   "20_TANKS_IP_DATA_RIO_07_FIRST_TANK_USD_FLOW" : Real = PLC "20_TANKS_IP_DATA".RIO_07.FIRST_TANK.USD_FLOW, 1 s
   "20_TANKS_IP_DATA_RIO_07_FIRST_TANK_MBG_FLOW" : Real = PLC "20_TANKS_IP_DATA".RIO_07.FIRST_TANK.MBG_FLOW, 1 s
   "504_Tank Grouping_DB2020_RUN TANK 14" : Bool = PLC "504_Tank Grouping_DB2020"."RUN TANK 14", 1 s
   "504_Tank Grouping_DB2020_RUN TANK 6" : Bool = PLC "504_Tank Grouping_DB2020"."RUN TANK 6", 1 s
   "504_Tank Grouping_DB2020_RUN TANK 8" : Bool = PLC "504_Tank Grouping_DB2020"."RUN TANK 8", 1 s
   "504_Tank Grouping_DB2020_RUN TANK 9" : Bool = PLC "504_Tank Grouping_DB2020"."RUN TANK 9", 1 s
   "504_Tank Grouping_DB2020_RUN TANK 10" : Bool = PLC "504_Tank Grouping_DB2020"."RUN TANK 10", 1 s
   "504_Tank Grouping_DB2020_RUN TANK 11" : Bool = PLC "504_Tank Grouping_DB2020"."RUN TANK 11", 1 s
   "504_Tank Grouping_DB2020_RUN TANK 12" : Bool = PLC "504_Tank Grouping_DB2020"."RUN TANK 12", 1 s
   "504_Tank Grouping_DB2020_RUN TANK 13" : Bool = PLC "504_Tank Grouping_DB2020"."RUN TANK 13", 1 s
   "504_Tank Grouping_DB2020_Sequence Time m Offset" : Time = PLC "504_Tank Grouping_DB2020"."Sequence Time m Offset", 1 s
   "20_TANKS_IP_DATA_RIO_01_FIRST_TANK_TANKS_PRESS" : Real = PLC "20_TANKS_IP_DATA".RIO_01.FIRST_TANK.TANKS_PRESS, 1 s
   "20_TANKS_IP_DATA_RIO_01_FIRST_TANK_BWT_LEVEL" : Real = PLC "20_TANKS_IP_DATA".RIO_01.FIRST_TANK.BWT_LEVEL, 1 s
   "20_TANKS_IP_DATA_RIO_01_FIRST_TANK_BWT_PH" : Real = PLC "20_TANKS_IP_DATA".RIO_01.FIRST_TANK.BWT_PH, 1 s
   "20_TANKS_IP_DATA_RIO_01_FIRST_TANK_BWT_DO" : Real = PLC "20_TANKS_IP_DATA".RIO_01.FIRST_TANK.BWT_DO, 1 s
   "20_TANKS_IP_DATA_RIO_01_FIRST_TANK_BWT_TEMP" : Real = PLC "20_TANKS_IP_DATA".RIO_01.FIRST_TANK.BWT_TEMP, 1 s
   "504_Tank Grouping_DB2020_Tank1 Min Time_ET" : Time = PLC "504_Tank Grouping_DB2020"."Tank1 Min Time".ET, 1 s
   "504_Tank Grouping_DB2020_Tank2 Min Time_ET" : Time = PLC "504_Tank Grouping_DB2020"."Tank2 Min Time".ET, 1 s
   "20_TANKS_IP_DATA_RIO_01_SECOND_TANK_TANKS_PRESS" : Real = PLC "20_TANKS_IP_DATA".RIO_01.SECOND_TANK.TANKS_PRESS, 1 s
   "20_TANKS_IP_DATA_RIO_01_SECOND_TANK_BWT_LEVEL" : Real = PLC "20_TANKS_IP_DATA".RIO_01.SECOND_TANK.BWT_LEVEL, 1 s
   "20_TANKS_IP_DATA_RIO_01_SECOND_TANK_BWT_PH" : Real = PLC "20_TANKS_IP_DATA".RIO_01.SECOND_TANK.BWT_PH, 1 s
   "20_TANKS_IP_DATA_RIO_01_SECOND_TANK_BWT_DO" : Real = PLC "20_TANKS_IP_DATA".RIO_01.SECOND_TANK.BWT_DO, 1 s
   "20_TANKS_IP_DATA_RIO_01_SECOND_TANK_BWT_TEMP" : Real = PLC "20_TANKS_IP_DATA".RIO_01.SECOND_TANK.BWT_TEMP, 1 s
   "20_TANKS_IP_DATA_RIO_01_THIRD_TANK_TANKS_PRESS" : Real = PLC "20_TANKS_IP_DATA".RIO_01.THIRD_TANK.TANKS_PRESS, 1 s
   "20_TANKS_IP_DATA_RIO_01_THIRD_TANK_BWT_LEVEL" : Real = PLC "20_TANKS_IP_DATA".RIO_01.THIRD_TANK.BWT_LEVEL, 1 s
   "20_TANKS_IP_DATA_RIO_01_THIRD_TANK_BWT_PH" : Real = PLC "20_TANKS_IP_DATA".RIO_01.THIRD_TANK.BWT_PH, 1 s
   "20_TANKS_IP_DATA_RIO_01_THIRD_TANK_BWT_DO" : Real = PLC "20_TANKS_IP_DATA".RIO_01.THIRD_TANK.BWT_DO, 1 s
   "20_TANKS_IP_DATA_RIO_01_THIRD_TANK_BWT_TEMP" : Real = PLC "20_TANKS_IP_DATA".RIO_01.THIRD_TANK.BWT_TEMP, 1 s
   "504_Tank Grouping_DB2020_Tank4 Min Time_ET" : Time = PLC "504_Tank Grouping_DB2020"."Tank4 Min Time".ET, 1 s
   "504_Tank Grouping_DB2020_Tank3 Min Time_ET" : Time = PLC "504_Tank Grouping_DB2020"."Tank3 Min Time".ET, 1 s
   "504_Tank Grouping_DB2020_Tank5 Min Time_ET" : Time = PLC "504_Tank Grouping_DB2020"."Tank5 Min Time".ET, 1 s
   "20_TANKS_IP_DATA_RIO_03_FIRST_TANK_TANKS_PRESS" : Real = PLC "20_TANKS_IP_DATA".RIO_03.FIRST_TANK.TANKS_PRESS, 1 s
   "20_TANKS_IP_DATA_RIO_03_FIRST_TANK_BWT_LEVEL" : Real = PLC "20_TANKS_IP_DATA".RIO_03.FIRST_TANK.BWT_LEVEL, 1 s
   "20_TANKS_IP_DATA_RIO_03_FIRST_TANK_BWT_PH" : Real = PLC "20_TANKS_IP_DATA".RIO_03.FIRST_TANK.BWT_PH, 1 s
   "20_TANKS_IP_DATA_RIO_03_FIRST_TANK_BWT_DO" : Real = PLC "20_TANKS_IP_DATA".RIO_03.FIRST_TANK.BWT_DO, 1 s
   "20_TANKS_IP_DATA_RIO_03_FIRST_TANK_BWT_TEMP" : Real = PLC "20_TANKS_IP_DATA".RIO_03.FIRST_TANK.BWT_TEMP, 1 s
   "504_Tank Grouping_DB2020_Tank6 Min Time_ET" : Time = PLC "504_Tank Grouping_DB2020"."Tank6 Min Time".ET, 1 s
   "20_TANKS_IP_DATA_RIO_03_SECOND_TANK_TANKS_PRESS" : Real = PLC "20_TANKS_IP_DATA".RIO_03.SECOND_TANK.TANKS_PRESS, 1 s
   "20_TANKS_IP_DATA_RIO_03_SECOND_TANK_BWT_LEVEL" : Real = PLC "20_TANKS_IP_DATA".RIO_03.SECOND_TANK.BWT_LEVEL, 1 s
   "20_TANKS_IP_DATA_RIO_03_SECOND_TANK_BWT_PH" : Real = PLC "20_TANKS_IP_DATA".RIO_03.SECOND_TANK.BWT_PH, 1 s
   "20_TANKS_IP_DATA_RIO_03_SECOND_TANK_BWT_DO" : Real = PLC "20_TANKS_IP_DATA".RIO_03.SECOND_TANK.BWT_DO, 1 s
   "20_TANKS_IP_DATA_RIO_03_SECOND_TANK_BWT_TEMP" : Real = PLC "20_TANKS_IP_DATA".RIO_03.SECOND_TANK.BWT_TEMP, 1 s
   "504_Tank Grouping_DB2020_Tank7 Min Time_ET" : Time = PLC "504_Tank Grouping_DB2020"."Tank7 Min Time".ET, 1 s
   "20_TANKS_IP_DATA_RIO_04_FIRST_TANK_TANKS_PRESS" : Real = PLC "20_TANKS_IP_DATA".RIO_04.FIRST_TANK.TANKS_PRESS, 1 s
   "20_TANKS_IP_DATA_RIO_04_FIRST_TANK_BWT_LEVEL" : Real = PLC "20_TANKS_IP_DATA".RIO_04.FIRST_TANK.BWT_LEVEL, 1 s
   "20_TANKS_IP_DATA_RIO_04_FIRST_TANK_BWT_PH" : Real = PLC "20_TANKS_IP_DATA".RIO_04.FIRST_TANK.BWT_PH, 1 s
   "20_TANKS_IP_DATA_RIO_04_FIRST_TANK_BWT_DO" : Real = PLC "20_TANKS_IP_DATA".RIO_04.FIRST_TANK.BWT_DO, 1 s
   "20_TANKS_IP_DATA_RIO_04_FIRST_TANK_BWT_TEMP" : Real = PLC "20_TANKS_IP_DATA".RIO_04.FIRST_TANK.BWT_TEMP, 1 s
   "504_Tank Grouping_DB2020_Tank8 Min Time_ET" : Time = PLC "504_Tank Grouping_DB2020"."Tank8 Min Time".ET, 1 s
   "20_TANKS_IP_DATA_RIO_04_SECOND_TANK_TANKS_PRESS" : Real = PLC "20_TANKS_IP_DATA".RIO_04.SECOND_TANK.TANKS_PRESS, 1 s
   "20_TANKS_IP_DATA_RIO_04_SECOND_TANK_BWT_LEVEL" : Real = PLC "20_TANKS_IP_DATA".RIO_04.SECOND_TANK.BWT_LEVEL, 1 s
   "20_TANKS_IP_DATA_RIO_04_SECOND_TANK_BWT_PH" : Real = PLC "20_TANKS_IP_DATA".RIO_04.SECOND_TANK.BWT_PH, 1 s
   "20_TANKS_IP_DATA_RIO_04_SECOND_TANK_BWT_DO" : Real = PLC "20_TANKS_IP_DATA".RIO_04.SECOND_TANK.BWT_DO, 1 s
   "20_TANKS_IP_DATA_RIO_04_SECOND_TANK_BWT_TEMP" : Real = PLC "20_TANKS_IP_DATA".RIO_04.SECOND_TANK.BWT_TEMP, 1 s
   "504_Tank Grouping_DB2020_Tank9 Min Time_ET" : Time = PLC "504_Tank Grouping_DB2020"."Tank9 Min Time".ET, 1 s
   "20_TANKS_IP_DATA_RIO_05_FIRST_TANK_TANKS_PRESS" : Real = PLC "20_TANKS_IP_DATA".RIO_05.FIRST_TANK.TANKS_PRESS, 1 s
   "20_TANKS_IP_DATA_RIO_05_FIRST_TANK_BWT_LEVEL" : Real = PLC "20_TANKS_IP_DATA".RIO_05.FIRST_TANK.BWT_LEVEL, 1 s
   "20_TANKS_IP_DATA_RIO_05_FIRST_TANK_BWT_PH" : Real = PLC "20_TANKS_IP_DATA".RIO_05.FIRST_TANK.BWT_PH, 1 s
   "20_TANKS_IP_DATA_RIO_05_FIRST_TANK_BWT_DO" : Real = PLC "20_TANKS_IP_DATA".RIO_05.FIRST_TANK.BWT_DO, 1 s
   "20_TANKS_IP_DATA_RIO_05_FIRST_TANK_BWT_TEMP" : Real = PLC "20_TANKS_IP_DATA".RIO_05.FIRST_TANK.BWT_TEMP, 1 s
   "504_Tank Grouping_DB2020_Tank10 Min Time_ET" : Time = PLC "504_Tank Grouping_DB2020"."Tank10 Min Time".ET, 1 s
   "20_TANKS_IP_DATA_RIO_05_SECOND_TANK_TANKS_PRESS" : Real = PLC "20_TANKS_IP_DATA".RIO_05.SECOND_TANK.TANKS_PRESS, 1 s
   "20_TANKS_IP_DATA_RIO_05_SECOND_TANK_BWT_LEVEL" : Real = PLC "20_TANKS_IP_DATA".RIO_05.SECOND_TANK.BWT_LEVEL, 1 s
   "20_TANKS_IP_DATA_RIO_05_SECOND_TANK_BWT_PH" : Real = PLC "20_TANKS_IP_DATA".RIO_05.SECOND_TANK.BWT_PH, 1 s
   "20_TANKS_IP_DATA_RIO_05_SECOND_TANK_BWT_DO" : Real = PLC "20_TANKS_IP_DATA".RIO_05.SECOND_TANK.BWT_DO, 1 s
   "20_TANKS_IP_DATA_RIO_05_SECOND_TANK_BWT_TEMP" : Real = PLC "20_TANKS_IP_DATA".RIO_05.SECOND_TANK.BWT_TEMP, 1 s
   "20_TANKS_IP_DATA_RIO_06_FIRST_TANK_TANKS_PRESS" : Real = PLC "20_TANKS_IP_DATA".RIO_06.FIRST_TANK.TANKS_PRESS, 1 s
   "20_TANKS_IP_DATA_RIO_06_FIRST_TANK_BWT_LEVEL" : Real = PLC "20_TANKS_IP_DATA".RIO_06.FIRST_TANK.BWT_LEVEL, 1 s
   "20_TANKS_IP_DATA_RIO_06_FIRST_TANK_BWT_PH" : Real = PLC "20_TANKS_IP_DATA".RIO_06.FIRST_TANK.BWT_PH, 1 s
   "20_TANKS_IP_DATA_RIO_06_FIRST_TANK_BWT_DO" : Real = PLC "20_TANKS_IP_DATA".RIO_06.FIRST_TANK.BWT_DO, 1 s
   "20_TANKS_IP_DATA_RIO_06_FIRST_TANK_BWT_TEMP" : Real = PLC "20_TANKS_IP_DATA".RIO_06.FIRST_TANK.BWT_TEMP, 1 s
   "504_Tank Grouping_DB2020_Tank12 Min Time_ET" : Time = PLC "504_Tank Grouping_DB2020"."Tank12 Min Time".ET, 1 s
   "20_TANKS_IP_DATA_RIO_06_SECOND_TANK_TANKS_PRESS" : Real = PLC "20_TANKS_IP_DATA".RIO_06.SECOND_TANK.TANKS_PRESS, 1 s
   "20_TANKS_IP_DATA_RIO_06_SECOND_TANK_BWT_LEVEL" : Real = PLC "20_TANKS_IP_DATA".RIO_06.SECOND_TANK.BWT_LEVEL, 1 s
   "20_TANKS_IP_DATA_RIO_06_SECOND_TANK_BWT_PH" : Real = PLC "20_TANKS_IP_DATA".RIO_06.SECOND_TANK.BWT_PH, 1 s
   "20_TANKS_IP_DATA_RIO_06_SECOND_TANK_BWT_DO" : Real = PLC "20_TANKS_IP_DATA".RIO_06.SECOND_TANK.BWT_DO, 1 s
   "20_TANKS_IP_DATA_RIO_06_SECOND_TANK_BWT_TEMP" : Real = PLC "20_TANKS_IP_DATA".RIO_06.SECOND_TANK.BWT_TEMP, 1 s
   "504_Tank Grouping_DB2020_Tank13 Min Time_ET" : Time = PLC "504_Tank Grouping_DB2020"."Tank13 Min Time".ET, 1 s
   "504_Tank Grouping_DB2020_Tank14 Min Time_ET" : Time = PLC "504_Tank Grouping_DB2020"."Tank14 Min Time".ET, 1 s
   "20_TANKS_IP_DATA_RIO_07_FIRST_TANK_TANKS_PRESS" : Real = PLC "20_TANKS_IP_DATA".RIO_07.FIRST_TANK.TANKS_PRESS, 1 s
   "20_TANKS_IP_DATA_RIO_07_FIRST_TANK_BWT_LEVEL" : Real = PLC "20_TANKS_IP_DATA".RIO_07.FIRST_TANK.BWT_LEVEL, 1 s
   "20_TANKS_IP_DATA_RIO_07_FIRST_TANK_BWT_PH" : Real = PLC "20_TANKS_IP_DATA".RIO_07.FIRST_TANK.BWT_PH, 1 s
   "20_TANKS_IP_DATA_RIO_07_FIRST_TANK_BWT_DO" : Real = PLC "20_TANKS_IP_DATA".RIO_07.FIRST_TANK.BWT_DO, 1 s
   "20_TANKS_IP_DATA_RIO_07_FIRST_TANK_BWT_TEMP" : Real = PLC "20_TANKS_IP_DATA".RIO_07.FIRST_TANK.BWT_TEMP, 1 s
   "504_Tank Grouping_DB2020_RUN" : Bool = PLC "504_Tank Grouping_DB2020".RUN, 1 s
   "80_From_HMI_Test Tank Request" : Bool = PLC "80_From_HMI".IGG_STND_ALN, 1 s
   "504_Tank Grouping_DB2020_Offset Timer_ET" : Time = PLC "504_Tank Grouping_DB2020"."Offset Timer".ET, 1 s
   "504_Tank Grouping_DB2020_Time Left Tank_Time Left Tank 7" : Real = PLC "504_Tank Grouping_DB2020"."Time Left Tank"."Time Left Tank 7", 1 s
   "504_Tank Grouping_DB2020_Time Left Tank_Time Left Tank 2" : Real = PLC "504_Tank Grouping_DB2020"."Time Left Tank"."Time Left Tank 2", 1 s
   "504_Tank Grouping_DB2020_Time Left Tank_Time Left Tank 3" : Real = PLC "504_Tank Grouping_DB2020"."Time Left Tank"."Time Left Tank 3", 1 s
   "504_Tank Grouping_DB2020_Time Left Tank_Time Left Tank 4" : Real = PLC "504_Tank Grouping_DB2020"."Time Left Tank"."Time Left Tank 4", 1 s
   "504_Tank Grouping_DB2020_Time Left Tank_Time Left Tank 5" : Real = PLC "504_Tank Grouping_DB2020"."Time Left Tank"."Time Left Tank 5", 1 s
   "504_Tank Grouping_DB2020_Time Left Tank_Time Left Tank 6" : Real = PLC "504_Tank Grouping_DB2020"."Time Left Tank"."Time Left Tank 6", 1 s
   "504_Tank Grouping_DB2020_Time Left Tank_Time Left Tank 8" : Real = PLC "504_Tank Grouping_DB2020"."Time Left Tank"."Time Left Tank 8", 1 s
   "504_Tank Grouping_DB2020_Time Left Tank_Time Left Tank 9" : Real = PLC "504_Tank Grouping_DB2020"."Time Left Tank"."Time Left Tank 9", 1 s
   "504_Tank Grouping_DB2020_Time Left Tank_Time Left Tank 10" : Real = PLC "504_Tank Grouping_DB2020"."Time Left Tank"."Time Left Tank 10", 1 s
   "504_Tank Grouping_DB2020_Time Left Tank_Time Left Tank 11" : Real = PLC "504_Tank Grouping_DB2020"."Time Left Tank"."Time Left Tank 11", 1 s
   "504_Tank Grouping_DB2020_Time Left Tank_Time Left Tank 12" : Real = PLC "504_Tank Grouping_DB2020"."Time Left Tank"."Time Left Tank 12", 1 s
   "504_Tank Grouping_DB2020_Time Left Tank_Time Left Tank 13" : Real = PLC "504_Tank Grouping_DB2020"."Time Left Tank"."Time Left Tank 13", 1 s
   "504_Tank Grouping_DB2020_Time Left Tank_Time Left Tank 14" : Real = PLC "504_Tank Grouping_DB2020"."Time Left Tank"."Time Left Tank 14", 1 s
   "504_Tank Grouping_DB2020_Time Left Tank_Time Left Tank 1" : Real = PLC "504_Tank Grouping_DB2020"."Time Left Tank"."Time Left Tank 1", 1 s
   "504_Tank Grouping_DB2020_SetGroupSR" : Bool = PLC "504_Tank Grouping_DB2020".SetGroupSR, 1 s
   "504_Tank Grouping_DB2020_Diff Time Remain" : DInt = PLC "504_Tank Grouping_DB2020"."Diff Time Remain", 1 s
   "2084_Setpoints_FIT417_LoLo" : Real = PLC "2084_Setpoints".FIT417_LoLo, 1 s
   "2084_Setpoints_FIT417_Lo" : Real = PLC "2084_Setpoints".FIT417_Lo, 1 s
   "2084_Setpoints_FIT417_Hi" : Real = PLC "2084_Setpoints".FIT417_Hi, 1 s
   "2084_Setpoints_FIT417_HiHi" : Real = PLC "2084_Setpoints".FIT417_HiHi, 1 s
   "2084_Setpoints_FIT419_LoLo" : Real = PLC "2084_Setpoints".FIT419_LoLo, 1 s
   "2084_Setpoints_FIT419_Lo" : Real = PLC "2084_Setpoints".FIT419_Lo, 1 s
   "2084_Setpoints_FIT419_Hi" : Real = PLC "2084_Setpoints".FIT419_Hi, 1 s
   "2084_Setpoints_FIT419_HiHi" : Real = PLC "20_TANKS_IP_DATA".RIO_02.FIRST_TANK.TANK_VENT_B_OPEN, 1 s
   "2084_Setpoints_LT421_Lo" : Real = PLC "2084_Setpoints".LT421_Lo, 1 s
   "2084_Setpoints_LT421_Hi" : Real = PLC "2084_Setpoints".LT421_Hi, 1 s
   "2084_Setpoints_TX426 Port PH Lo" : Real = PLC "2084_Setpoints"."TX426 Port PH Lo", 1 s
   "2084_Setpoints_TX426 Port PH High" : Real = PLC "2084_Setpoints"."TX426 Port PH High", 1 s
   "2084_Setpoints_TX428 Port DO Lo" : Real = PLC "2084_Setpoints"."TX428 Port DO Lo", 1 s
   "2084_Setpoints_TX428 Port DO High" : Real = PLC "2084_Setpoints"."TX428 Port DO High", 1 s
   "2084_Setpoints_TX425 Star PH Lo" : Real = PLC "2084_Setpoints"."TX425 Star PH Lo", 1 s
   "2084_Setpoints_TX425 Star PH High" : Real = PLC "2084_Setpoints"."TX425 Star PH High", 1 s
   "2084_Setpoints_TX427 Star DO Lo" : Real = PLC "2084_Setpoints"."TX427 Star DO Lo", 1 s
   "2084_Setpoints_TX427 Star DO High" : Real = PLC "2084_Setpoints"."TX427 Star DO High", 1 s
   "2084_Setpoints_Conf O2 Level Lo" : Real = PLC "2084_Setpoints"."Conf O2 Level Lo", 1 s
   "2084_Setpoints_Conf O2 Level Lo Lo" : Real = PLC "2084_Setpoints"."Conf O2 Level Lo Lo", 1 s
   "20_TANKS_IP_DATA_RIO_03_FIRST_TANK_O2_MONITOR" : Real = PLC FIT420_5P_ALM_ANALOG_DB."LOW LEVEL VALUE (L)", 1 s
   "20_TANKS_IP_DATA_RIO_03_SECOND_TANK_O2_MONITOR" : Real = PLC "20_TANKS_IP_DATA".RIO_03.SECOND_TANK.O2_MONITOR, 1 s
   "20_TANKS_IP_DATA_RIO_03_FIRST_TANK_DECK_IG_PRESS" : Real = PLC "20_TANKS_IP_DATA".RIO_03.FIRST_TANK.DECK_IG_PRESS, 1 s
   "20_TANKS_IP_DATA_RIO_01_THIRD_TANK_O2_MONITOR" : Real = PLC "20_TANKS_IP_DATA".RIO_01.THIRD_TANK.O2_MONITOR, 1 s
   "20_TANKS_IP_DATA_RIO_01_THIRD_TANK_DECK_IG_PRESS" : Real = PLC "20_TANKS_IP_DATA".RIO_01.THIRD_TANK.DECK_IG_PRESS, 1 s
   "20_TANKS_IP_DATA_RIO_01_FIRST_TANK_DECK_IG_PRESS" : Real = PLC "20_TANKS_IP_DATA".RIO_01.FIRST_TANK.DECK_IG_PRESS, 1 s
   "20_TANKS_IP_DATA_RIO_01_FIRST_TANK_O2_MONITOR" : Real = PLC "20_TANKS_IP_DATA".RIO_01.FIRST_TANK.O2_MONITOR, 1 s
   "20_TANKS_IP_DATA_RIO_04_FIRST_TANK_DECK_IG_PRESS" : Real = PLC "20_TANKS_IP_DATA".RIO_04.FIRST_TANK.DECK_IG_PRESS, 1 s
   "20_TANKS_IP_DATA_RIO_04_FIRST_TANK_O2_MONITOR" : Real = PLC "20_TANKS_IP_DATA".RIO_04.FIRST_TANK.O2_MONITOR, 1 s
   "20_TANKS_IP_DATA_RIO_04_SECOND_TANK_O2_MONITOR" : Real = PLC "20_TANKS_IP_DATA".RIO_04.SECOND_TANK.O2_MONITOR, 1 s
   "20_TANKS_IP_DATA_RIO_05_FIRST_TANK_DECK_IG_PRESS" : Real = PLC "20_TANKS_IP_DATA".RIO_05.FIRST_TANK.DECK_IG_PRESS, 1 s
   "20_TANKS_IP_DATA_RIO_05_FIRST_TANK_O2_MONITOR" : Real = PLC "20_TANKS_IP_DATA".RIO_05.FIRST_TANK.O2_MONITOR, 1 s
   "20_TANKS_IP_DATA_RIO_05_SECOND_TANK_O2_MONITOR" : Real = PLC "20_TANKS_IP_DATA".RIO_05.SECOND_TANK.O2_MONITOR, 1 s
   "20_TANKS_IP_DATA_RIO_06_FIRST_TANK_DECK_IG_PRESS" : Real = PLC "20_TANKS_IP_DATA".RIO_06.FIRST_TANK.DECK_IG_PRESS, 1 s
   "20_TANKS_IP_DATA_RIO_06_FIRST_TANK_O2_MONITOR" : Real = PLC "20_TANKS_IP_DATA".RIO_06.FIRST_TANK.O2_MONITOR, 1 s
   "20_TANKS_IP_DATA_RIO_07_FIRST_TANK_O2_MONITOR" : Real = PLC "10_DI_DATA".P_304_ENBLD, 1 s
   "20_TANKS_IP_DATA_RIO_07_FIRST_TANK_DECK_IG_PRESS" : Real = PLC "20_TANKS_IP_DATA".RIO_07.FIRST_TANK.DECK_IG_PRESS, 1 s
   "2062_Warning_Data_BTCS_WARNING_WORD_09" : Word = PLC "2062_Warning_Data".BTCS_WARNING_WORD_09 AT %DB2062.DBW16, 1 s
   "2086_Times_Tank Alarm Reset Time" : Time = PLC "2086_Times"."Tank Alarm Reset Time", 1 s
   "2086_Times_Alarm Enable Delay" : Time = PLC "2086_Times"."Alarm Enable Delay", 1 s
   "2062_Warning_Data_BTCS_WARNING_WORD_10" : Word = PLC "2062_Warning_Data".BTCS_WARNING_WORD_10 AT %DB2062.DBW18, 1 s
   "2062_Warning_Data_BTCS_WARNING_WORD_11" : Word = PLC "2062_Warning_Data".BTCS_WARNING_WORD_11 AT %DB2062.DBW20, 1 s
   "LT422 FPT  TANK LEVEL ALARM_LOW LEVEL VALUE (L)" : Real = PLC "LT422 FPT  TANK LEVEL ALARM"."LOW LEVEL VALUE (L)" AT %DB2226.DBD26, 1 s
   "LT422 FPT  TANK LEVEL ALARM_ALARM L" : Bool = PLC "LT422 FPT  TANK LEVEL ALARM"."ALARM L" AT %DB2226.DBX48.2, 1 s
   "2062_Warning_Data_Alarm Tank FPT" : Bool = PLC "2062_Warning_Data"."Alarm Tank FPT" AT %DB2062.DBX22.1, 1 s
   "2062_Warning_Data_Water Level Override FPT" : Bool = PLC "2062_Warning_Data"."Water Level Override FPT" AT %DB2062.DBX360.0, 1 s
   "LT422 1P  TANK LEVEL ALARM_ALARM L" : Bool = PLC "LT422 1P  TANK LEVEL ALARM"."ALARM L" AT %DB2227.DBX48.2, 1 s
   "2062_Warning_Data_Alarm Tank P1" : Bool = PLC "2062_Warning_Data"."Alarm Tank P1" AT %DB2062.DBX22.2, 1 s
   "2062_Warning_Data_Water Level Override 1P" : Bool = PLC "2062_Warning_Data"."Water Level Override 1P" AT %DB2062.DBX360.1, 1 s
   "LT421 1S  TANK LEVEL ALARM_ALARM L" : Bool = PLC "LT421 1S  TANK LEVEL ALARM"."ALARM L" AT %DB2228.DBX48.2, 1 s
   "2062_Warning_Data_Alarm Tank S1" : Bool = PLC "2062_Warning_Data"."Alarm Tank S1" AT %DB2062.DBX22.3, 1 s
   "FIT418_2P_ALM_ANALOG_DB_ALARM L" : Bool = PLC FIT418_2P_ALM_ANALOG_DB."ALARM L" AT %DB2064.DBX48.2, 1 s
   "2062_Warning_Data_Alarm Tank P2" : Bool = PLC "2062_Warning_Data"."Alarm Tank P2" AT %DB2062.DBX22.4, 1 s
   "2062_Warning_Data_Water Level Override 2P" : Bool = PLC "2062_Warning_Data"."Water Level Override 2P" AT %DB2062.DBX360.3, 1 s
   "2062_Warning_Data_Water Level Override 1S" : Bool = PLC "2062_Warning_Data"."Water Level Override 1S" AT %DB2062.DBX360.2, 1 s
   "LT421 2S  TANK LEVEL ALARM_ALARM L" : Bool = PLC "LT421 2S  TANK LEVEL ALARM"."ALARM L" AT %DB2230.DBX48.2, 1 s
   "2062_Warning_Data_Alarm Tank S2" : Bool = PLC "2062_Warning_Data"."Alarm Tank S2" AT %DB2062.DBX22.5, 1 s
   "2062_Warning_Data_Water Level Override 2S" : Bool = PLC "2062_Warning_Data"."Water Level Override 2S" AT %DB2062.DBX360.4, 1 s
   "LT422 3P  TANK LEVEL ALARM_ALARM L" : Bool = PLC "LT422 3P  TANK LEVEL ALARM"."ALARM L" AT %DB2231.DBX48.2, 1 s
   "2062_Warning_Data_Alarm Tank P3" : Bool = PLC "2062_Warning_Data"."Alarm Tank P3" AT %DB2062.DBX22.6, 1 s
   "2062_Warning_Data_Water Level Override 3P" : Bool = PLC "2062_Warning_Data"."Water Level Override 3P" AT %DB2062.DBX360.5, 1 s
   "LT421 3S  TANK LEVEL ALARM_ALARM L" : Bool = PLC "LT421 3S  TANK LEVEL ALARM"."ALARM L" AT %DB2232.DBX48.2, 1 s
   "2062_Warning_Data_Alarm Tank S3" : Bool = PLC "2062_Warning_Data"."Alarm Tank S3" AT %DB2062.DBX22.7, 1 s
   "2062_Warning_Data_Water Level Override 3S" : Bool = PLC "2062_Warning_Data"."Water Level Override 3S" AT %DB2062.DBX360.6, 1 s
   "LT422 4P  TANK LEVEL ALARM_ALARM L" : Bool = PLC "LT422 4P  TANK LEVEL ALARM"."ALARM L" AT %DB2233.DBX48.2, 1 s
   "2062_Warning_Data_Alarm Tank P4" : Bool = PLC "2062_Warning_Data"."Alarm Tank P4" AT %DB2062.DBX23.0, 1 s
   "2062_Warning_Data_Water Level Override 4P" : Bool = PLC "2062_Warning_Data"."Water Level Override 4P" AT %DB2062.DBX360.7, 1 s
   "LT421 4S  TANK LEVEL ALARM_ALARM L" : Bool = PLC "LT421 4S  TANK LEVEL ALARM"."ALARM L" AT %DB2234.DBX48.2, 1 s
   "2062_Warning_Data_Alarm Tank S4" : Bool = PLC "2062_Warning_Data"."Alarm Tank S4" AT %DB2062.DBX23.1, 1 s
   "2062_Warning_Data_Water Level Override 4S" : Bool = PLC "2062_Warning_Data"."Water Level Override 4S" AT %DB2062.DBX361.0, 1 s
   "LT422 5P  TANK LEVEL ALARM_ALARM L" : Bool = PLC "LT422 5P  TANK LEVEL ALARM"."ALARM L" AT %DB2235.DBX48.2, 1 s
   "2062_Warning_Data_Alarm Tank P5" : Bool = PLC "2062_Warning_Data"."Alarm Tank P5" AT %DB2062.DBX23.2, 1 s
   "2062_Warning_Data_Water Level Override 5P" : Bool = PLC "2062_Warning_Data"."Water Level Override 5P" AT %DB2062.DBX361.1, 1 s
   "LT421 5S  TANK LEVEL ALARM_ALARM L" : Bool = PLC "LT421 5S  TANK LEVEL ALARM"."ALARM L" AT %DB2236.DBX48.2, 1 s
   "2062_Warning_Data_Alarm Tank S5" : Bool = PLC "2062_Warning_Data"."Alarm Tank S5" AT %DB2062.DBX23.3, 1 s
   "2062_Warning_Data_Water Level Override 5S" : Bool = PLC "2062_Warning_Data"."Water Level Override 5S" AT %DB2062.DBX361.2, 1 s
   "LT422 6P  TANK LEVEL ALARM_ALARM L" : Bool = PLC "LT422 6P  TANK LEVEL ALARM"."ALARM L" AT %DB2237.DBX48.2, 1 s
   "2062_Warning_Data_Alarm Tank P6" : Bool = PLC "2062_Warning_Data"."Alarm Tank P6" AT %DB2062.DBX23.4, 1 s
   "2062_Warning_Data_Water Level Override 6P" : Bool = PLC "2062_Warning_Data"."Water Level Override 6P" AT %DB2062.DBX361.3, 1 s
   "LT421 6S  TANK LEVEL ALARM_ALARM L" : Bool = PLC "LT421 6S  TANK LEVEL ALARM"."ALARM L" AT %DB2238.DBX48.2, 1 s
   "2062_Warning_Data_Alarm Tank S6" : Bool = PLC "2062_Warning_Data"."Alarm Tank S6" AT %DB2062.DBX23.5, 1 s
   "2062_Warning_Data_Water Level Override 6S" : Bool = PLC "2062_Warning_Data"."Water Level Override 6S" AT %DB2062.DBX361.4, 1 s
   "LT422 APT  TANK LEVEL ALARM_ALARM L" : Bool = PLC "LT422 APT  TANK LEVEL ALARM"."ALARM L" AT %DB2239.DBX48.2, 1 s
   "2062_Warning_Data_Alarm Tank APT" : Bool = PLC "2062_Warning_Data"."Alarm Tank APT" AT %DB2062.DBX23.6, 1 s
   "2062_Warning_Data_Water Level Override APT" : Bool = PLC "2062_Warning_Data"."Water Level Override APT" AT %DB2062.DBX361.5, 1 s
   "FPT GTT Isolation Valve Feedback - Opened" : Bool = PLC "FPT GTT Isolation Valve Feedback - Opened" AT %I0.0, 1 s
   "FPT GTT Isolation Valve Feedback - Closed" : Bool = PLC "FPT GTT Isolation Valve Feedback - Closed" AT %I0.1, 1 s
   "FPT Tank Vent Valve 1 Feedback - Opened" : Bool = PLC "FPT Tank Vent Valve 1 Feedback - Opened" AT %I0.2, 1 s
   "FPT Tank Vent Valve 1 Feedback - Closed" : Bool = PLC "FPT Tank Vent Valve 1 Feedback - Closed" AT %I0.3, 1 s
   "FPT Tank Vent Valve 2 Feedback - Opened" : Bool = PLC "FPT Tank Vent Valve 2 Feedback - Opened" AT %I0.4, 1 s
   "FPT Tank Vent Valve 2 Feedback - Closed" : Bool = PLC "FPT Tank Vent Valve 2 Feedback - Closed" AT %I0.5, 1 s
   "RIO1_SPR_DI_0_6" : Bool = PLC RIO1_SPR_DI_0_6 AT %I0.6, 1 s
   "RIO1_SPR_DI_0_7" : Bool = PLC RIO1_SPR_DI_0_7 AT %I0.7, 1 s
   "Tank 1P GTT Isolation Valve Feedback - Opened" : Bool = PLC "Tank 1P GTT Isolation Valve Feedback - Opened" AT %I3.0, 1 s
   "Tank 1P GTT Isolation Valve Feedback - Closed" : Bool = PLC "Tank 1P GTT Isolation Valve Feedback - Closed" AT %I3.1, 1 s
   "Tank 1P Tank Vent Valve 1 Feedback - Opened" : Bool = PLC "Tank 1P Tank Vent Valve 1 Feedback - Opened" AT %I3.2, 1 s
   "Tank 1P Tank Vent Valve 1 Feedback - Closed" : Bool = PLC "Tank 1P Tank Vent Valve 1 Feedback - Closed" AT %I3.3, 1 s
   "Tank 1P Tank Vent Valve 2 Feedback - Opened" : Bool = PLC "Tank 1P Tank Vent Valve 2 Feedback - Opened" AT %I3.4, 1 s
   "Tank 1P Tank Vent Valve 2 Feedback - Closed" : Bool = PLC "Tank 1P Tank Vent Valve 2 Feedback - Closed" AT %I3.5, 1 s
   "RIO1_SPR_DI_3_6" : Bool = PLC RIO1_SPR_DI_3_6 AT %I3.6, 1 s
   "RIO1_SPR_DI_3_7" : Bool = PLC RIO1_SPR_DI_3_7 AT %I3.7, 1 s
   "Tank 1S GTT Isolation Valve Feedback - Opened" : Bool = PLC "Tank 1S GTT Isolation Valve Feedback - Opened" AT %I6.0, 1 s
   "Tank 1S GTT Isolation Valve Feedback - Closed" : Bool = PLC "Tank 1S GTT Isolation Valve Feedback - Closed" AT %I6.1, 1 s
   "Tank 1S Tank Vent Valve 1 Feedback - Opened" : Bool = PLC "Tank 1S Tank Vent Valve 1 Feedback - Opened" AT %I6.2, 1 s
   "Tank 1S Tank Vent Valve 1 Feedback - Closed" : Bool = PLC "Tank 1S Tank Vent Valve 1 Feedback - Closed" AT %I6.3, 1 s
   "Tank 1S Tank Vent Valve 2 Feedback - Opened" : Bool = PLC "Tank 1S Tank Vent Valve 2 Feedback - Opened" AT %I6.4, 1 s
   "Tank 1S Tank Vent Valve 2 Feedback - Closed" : Bool = PLC "Tank 1S Tank Vent Valve 2 Feedback - Closed" AT %I6.5, 1 s
   "RIO1_SPR_DI_6_6" : Bool = PLC RIO1_SPR_DI_6_6 AT %I6.6, 1 s
   "RIO1_SPR_DI_6_7" : Bool = PLC RIO1_SPR_DI_6_7 AT %I6.7, 1 s
   "FPT BWT Level High High Switch" : Bool = PLC "FPT BWT Level High High Switch" AT %I9.0, 1 s
   "RIO1 Tanks Pressure Switch Hi Hi" : Bool = PLC "RIO1 Tanks Pressure Switch Hi Hi" AT %I9.1, 1 s
   "Tank 1P BWT Level High High Switch" : Bool = PLC "Tank 1P BWT Level High High Switch" AT %I9.2, 1 s
   "Tank 1S BWT Level High High Switch" : Bool = PLC "Tank 1S BWT Level High High Switch" AT %I9.3, 1 s
   "RIO1_SPR_DI_9_4" : Bool = PLC RIO1_SPR_DI_9_4 AT %I9.4, 1 s
   "RIO1_SPR_DI_9_5" : Bool = PLC RIO1_SPR_DI_9_5 AT %I9.5, 1 s
   "RIO1_SPR_DI_9_6" : Bool = PLC RIO1_SPR_DI_9_6 AT %I9.6, 1 s
   "RIO1_SPR_DI_9_7" : Bool = PLC RIO1_SPR_DI_9_7 AT %I9.7, 1 s
   "Tank 2P GTT Isolation Valve Feedback - Opened" : Bool = PLC "Tank 2P GTT Isolation Valve Feedback - Opened" AT %I15.0, 1 s
   "Tank 2P GTT Isolation Valve Feedback - Closed" : Bool = PLC "Tank 2P GTT Isolation Valve Feedback - Closed" AT %I15.1, 1 s
   "Tank 2P Tank Vent Valve 1 Feedback - Opened" : Bool = PLC "Tank 2P Tank Vent Valve 1 Feedback - Opened" AT %I15.2, 1 s
   "Tank 2P Tank Vent Valve 1 Feedback - Closed" : Bool = PLC "Tank 2P Tank Vent Valve 1 Feedback - Closed" AT %I15.3, 1 s
   "Tank 2P Tank Vent Valve 2 Feedback - Opened" : Bool = PLC "Tank 2P Tank Vent Valve 2 Feedback - Opened" AT %I15.4, 1 s
   "Tank 2P Tank Vent Valve 2 Feedback - Closed" : Bool = PLC "Tank 2P Tank Vent Valve 2 Feedback - Closed" AT %I15.5, 1 s
   "RIO2_SPR_DI_15_6" : Bool = PLC RIO2_SPR_DI_15_6 AT %I15.6, 1 s
   "RIO2_SPR_DI_15_7" : Bool = PLC RIO2_SPR_DI_15_7 AT %I15.7, 1 s
   "Tank 2S GTT Isolation Valve Feedback - Opened" : Bool = PLC "Tank 2S GTT Isolation Valve Feedback - Opened" AT %I18.0, 1 s
   "Tank 2S GTT Isolation Valve Feedback - Closed" : Bool = PLC "Tank 2S GTT Isolation Valve Feedback - Closed" AT %I18.1, 1 s
   "Tank 2S Tank Vent Valve 1 Feedback - Opened" : Bool = PLC "Tank 2S Tank Vent Valve 1 Feedback - Opened" AT %I18.2, 1 s
   "Tank 2S Tank Vent Valve 1 Feedback - Closed" : Bool = PLC "Tank 2S Tank Vent Valve 1 Feedback - Closed" AT %I18.3, 1 s
   "Tank 2S Tank Vent Valve 2 Feedback - Opened" : Bool = PLC "Tank 2S Tank Vent Valve 2 Feedback - Opened" AT %I18.4, 1 s
   "Tank 2S Tank Vent Valve 2 Feedback - Closed" : Bool = PLC "Tank 2S Tank Vent Valve 2 Feedback - Closed" AT %I18.5, 1 s
   "RIO2_SPR_DI_18_6" : Bool = PLC RIO2_SPR_DI_18_6 AT %I18.6, 1 s
   "RIO2_SPR_DI_18_7" : Bool = PLC RIO2_SPR_DI_18_7 AT %I18.7, 1 s
   "Tank 2P BWT Level High High Switch" : Bool = PLC "Tank 2P BWT Level High High Switch" AT %I21.0, 1 s
   "RIO2 Tanks Pressure Switch Hi Hi" : Bool = PLC "RIO2 Tanks Pressure Switch Hi Hi" AT %I21.1, 1 s
   "Tank 2S BWT Level High High Switch" : Bool = PLC "Tank 2S BWT Level High High Switch" AT %I21.2, 1 s
   "RIO2_SPR_DI_21_3" : Bool = PLC RIO2_SPR_DI_21_3 AT %I21.3, 1 s
   "RIO2_SPR_DI_21_4" : Bool = PLC RIO2_SPR_DI_21_4 AT %I21.4, 1 s
   "RIO2_SPR_DI_21_5" : Bool = PLC RIO2_SPR_DI_21_5 AT %I21.5, 1 s
   "RIO2_SPR_DI_21_6" : Bool = PLC RIO2_SPR_DI_21_6 AT %I21.6, 1 s
   "RIO2_SPR_DI_21_7" : Bool = PLC RIO2_SPR_DI_21_7 AT %I21.7, 1 s
   "Tank 3P GTT Isolation Valve Feedback - Opened" : Bool = PLC "Tank 3P GTT Isolation Valve Feedback - Opened" AT %I27.0, 1 s
   "Tank 3P GTT Isolation Valve Feedback - Closed" : Bool = PLC "Tank 3P GTT Isolation Valve Feedback - Closed" AT %I27.1, 1 s
   "Tank 3P Tank Vent Valve 1 Feedback - Opened" : Bool = PLC "Tank 3P Tank Vent Valve 1 Feedback - Opened" AT %I27.2, 1 s
   "Tank 3P Tank Vent Valve 1 Feedback - Closed" : Bool = PLC "Tank 3P Tank Vent Valve 1 Feedback - Closed" AT %I27.3, 1 s
   "Tank 3P Tank Vent Valve 2 Feedback - Opened" : Bool = PLC "Tank 3P Tank Vent Valve 2 Feedback - Opened" AT %I27.4, 1 s
   "Tank 3P Tank Vent Valve 2 Feedback - Closed" : Bool = PLC "Tank 3P Tank Vent Valve 2 Feedback - Closed" AT %I27.5, 1 s
   "RIO3_SPR_DI_27_6" : Bool = PLC RIO3_SPR_DI_27_6 AT %I27.6, 1 s
   "RIO3_SPR_DI_27_7" : Bool = PLC RIO3_SPR_DI_27_7 AT %I27.7, 1 s
   "Tank 3S GTT Isolation Valve Feedback - Opened" : Bool = PLC "Tank 3S GTT Isolation Valve Feedback - Opened" AT %I30.0, 1 s
   "Tank 3S GTT Isolation Valve Feedback - Closed" : Bool = PLC "Tank 3S GTT Isolation Valve Feedback - Closed" AT %I30.1, 1 s
   "Tank 3S Tank Vent Valve 1 Feedback - Opened" : Bool = PLC "Tank 3S Tank Vent Valve 1 Feedback - Opened" AT %I30.2, 1 s
   "Tank 3S Tank Vent Valve 1 Feedback - Closed" : Bool = PLC "Tank 3S Tank Vent Valve 1 Feedback - Closed" AT %I30.3, 1 s
   "Tank 3S Tank Vent Valve 2 Feedback - Opened" : Bool = PLC "Tank 3S Tank Vent Valve 2 Feedback - Opened" AT %I30.4, 1 s
   "Tank 3S Tank Vent Valve 2 Feedback - Closed" : Bool = PLC "Tank 3S Tank Vent Valve 2 Feedback - Closed" AT %I30.5, 1 s
   "RIO3_SPR_DI_30_6" : Bool = PLC RIO3_SPR_DI_30_6 AT %I30.6, 1 s
   "RIO3_SPR_DI_30_7" : Bool = PLC RIO3_SPR_DI_30_7 AT %I30.7, 1 s
   "Tank 3P BWT Level High High Switch" : Bool = PLC "Tank 3P BWT Level High High Switch" AT %I33.0, 1 s
   "RIO3 Tanks Pressure Switch Hi Hi" : Bool = PLC "RIO3 Tanks Pressure Switch Hi Hi" AT %I33.1, 1 s
   "Tank 3S BWT Level High High Switch" : Bool = PLC "Tank 3S BWT Level High High Switch" AT %I33.2, 1 s
   "RIO3_SPR_DI_33_3" : Bool = PLC RIO3_SPR_DI_33_3 AT %I33.3, 1 s
   "RIO3_SPR_DI_33_4" : Bool = PLC RIO3_SPR_DI_33_4 AT %I33.4, 1 s
   "RIO3_SPR_DI_33_5" : Bool = PLC RIO3_SPR_DI_33_5 AT %I33.5, 1 s
   "RIO3_SPR_DI_33_6" : Bool = PLC RIO3_SPR_DI_33_6 AT %I33.6, 1 s
   "RIO3_SPR_DI_33_7" : Bool = PLC RIO3_SPR_DI_33_7 AT %I33.7, 1 s
   "Tank 4P GTT Isolation Valve Feedback - Opened" : Bool = PLC "Tank 4P GTT Isolation Valve Feedback - Opened" AT %I39.0, 1 s
   "Tank 4P GTT Isolation Valve Feedback - Closed" : Bool = PLC "Tank 4P GTT Isolation Valve Feedback - Closed" AT %I39.1, 1 s
   "Tank 4P Tank Vent Valve 1 Feedback - Opened" : Bool = PLC "Tank 4P Tank Vent Valve 1 Feedback - Opened" AT %I39.2, 1 s
   "Tank 4P Tank Vent Valve 1 Feedback - Closed" : Bool = PLC "Tank 4P Tank Vent Valve 1 Feedback - Closed" AT %I39.3, 1 s
   "Tank 4P Tank Vent Valve 2 Feedback - Opened" : Bool = PLC "Tank 4P Tank Vent Valve 2 Feedback - Opened" AT %I39.4, 1 s
   "Tank 4P Tank Vent Valve 2 Feedback - Closed" : Bool = PLC "Tank 4P Tank Vent Valve 2 Feedback - Closed" AT %I39.5, 1 s
   "RIO4_SPR_DI_139_6" : Bool = PLC RIO4_SPR_DI_139_6 AT %I39.6, 1 s
   "RIO4_SPR_DI_139_7" : Bool = PLC RIO4_SPR_DI_139_7 AT %I39.7, 1 s
   "Tank 4S GTT Isolation Valve Feedback - Opened" : Bool = PLC "Tank 4S GTT Isolation Valve Feedback - Opened" AT %I42.0, 1 s
   "Tank 4S GTT Isolation Valve Feedback - Closed" : Bool = PLC "Tank 4S GTT Isolation Valve Feedback - Closed" AT %I42.1, 1 s
   "Tank 4S Tank Vent Valve 1 Feedback - Opened" : Bool = PLC "Tank 4S Tank Vent Valve 1 Feedback - Opened" AT %I42.2, 1 s
   "Tank 4S Tank Vent Valve 1 Feedback - Closed" : Bool = PLC "Tank 4S Tank Vent Valve 1 Feedback - Closed" AT %I42.3, 1 s
   "Tank 4S Tank Vent Valve 2 Feedback - Opened" : Bool = PLC "Tank 4S Tank Vent Valve 2 Feedback - Opened" AT %I42.4, 1 s
   "Tank 4S Tank Vent Valve 2 Feedback - Closed" : Bool = PLC "Tank 4S Tank Vent Valve 2 Feedback - Closed" AT %I42.5, 1 s
   "RIO4_SPR_DI_142_6" : Bool = PLC RIO4_SPR_DI_142_6 AT %I42.6, 1 s
   "RIO4_SPR_DI_142_7" : Bool = PLC RIO4_SPR_DI_142_7 AT %I42.7, 1 s
   "Tank 4P BWT Level High High Switch" : Bool = PLC "Tank 4P BWT Level High High Switch" AT %I45.0, 1 s
   "RIO4 Tanks Pressure Switch Hi Hi" : Bool = PLC "RIO4 Tanks Pressure Switch Hi Hi" AT %I45.1, 1 s
   "Tank 4S BWT Level High High Switch" : Bool = PLC "Tank 4S BWT Level High High Switch" AT %I45.2, 1 s
   "RIO4_SPR_DI_145_3" : Bool = PLC RIO4_SPR_DI_145_3 AT %I45.3, 1 s
   "RIO4_SPR_DI_145_4" : Bool = PLC RIO4_SPR_DI_145_4 AT %I45.4, 1 s
   "RIO4_SPR_DI_145_5" : Bool = PLC RIO4_SPR_DI_145_5 AT %I45.5, 1 s
   "RIO4_SPR_DI_145_6" : Bool = PLC RIO4_SPR_DI_145_6 AT %I45.6, 1 s
   "RIO4_SPR_DI_145_7" : Bool = PLC RIO4_SPR_DI_145_7 AT %I45.7, 1 s
   "Tank 5P GTT Isolation Valve Feedback - Opened" : Bool = PLC "Tank 5P GTT Isolation Valve Feedback - Opened" AT %I51.0, 1 s
   "Tank 5P GTT Isolation Valve Feedback - Closed" : Bool = PLC "Tank 5P GTT Isolation Valve Feedback - Closed" AT %I51.1, 1 s
   "Tank 5P Tank Vent Valve 1 Feedback - Opened" : Bool = PLC "Tank 5P Tank Vent Valve 1 Feedback - Opened" AT %I51.2, 1 s
   "Tank 5P Tank Vent Valve 1 Feedback - Closed" : Bool = PLC "Tank 5P Tank Vent Valve 1 Feedback - Closed" AT %I51.3, 1 s
   "Tank 5P Tank Vent Valve 2 Feedback - Opened" : Bool = PLC "Tank 5P Tank Vent Valve 2 Feedback - Opened" AT %I51.4, 1 s
   "Tank 5P Tank Vent Valve 2 Feedback - Closed" : Bool = PLC "Tank 5P Tank Vent Valve 2 Feedback - Closed" AT %I51.5, 1 s
   "RIO5_SPR_DI_51_6" : Bool = PLC RIO5_SPR_DI_51_6 AT %I51.6, 1 s
   "RIO5_SPR_DI_51_7" : Bool = PLC RIO5_SPR_DI_51_7 AT %I51.7, 1 s
   "Tank 5S GTT Isolation Valve Feedback - Opened" : Bool = PLC "Tank 5S GTT Isolation Valve Feedback - Opened" AT %I54.0, 1 s
   "Tank 5S GTT Isolation Valve Feedback - Closed" : Bool = PLC "Tank 5S GTT Isolation Valve Feedback - Closed" AT %I54.1, 1 s
   "Tank 5S Tank Vent Valve 1 Feedback - Opened" : Bool = PLC "Tank 5S Tank Vent Valve 1 Feedback - Opened" AT %I54.2, 1 s
   "Tank 5S Tank Vent Valve 1 Feedback - Closed" : Bool = PLC "Tank 5S Tank Vent Valve 1 Feedback - Closed" AT %I54.3, 1 s
   "Tank 5S Tank Vent Valve 2 Feedback - Opened" : Bool = PLC "Tank 5S Tank Vent Valve 2 Feedback - Opened" AT %I54.4, 1 s